// TIA Portal project "Oshop-Demo_v2" (V16)

(* hardware
DEVICE "ET 200SP-Station_1"  ET 200SP-Station
   slot 0: "Baugruppenträger_0"  Rack  6ES5 710-8MAx1
   slot 1: "PLC_1"  CPU 1512SP-1 PN  6ES7 512-1DK01-0AB0  V2.1
      slot 32768: "PROFINET-Schnittstelle_1"  X1
   slot 2: "DI 8x24VDC HF_1"  DI 8x24VDC HF  6ES7 131-6BF00-0CA0  V2.0
      slot 1: "DI 8x24VDC HF_1"  DI 8x24VDC HF
   slot 3: "CM 4xIO-Link_1"  CM 4xIO-Link  6ES7 137-6BD00-0BA0  V2.2
      slot 1: "CM 4xIO-Link_1"  6ES7 137-6BD00-0BA0
   slot 4: "DQ 8x24VDC/0.5A HF_1"  DQ 8x24VDC/0.5A HF  6ES7 132-6BF00-0CA0  V2.0
      slot 1: "DQ 8x24VDC/0.5A HF_1"  DQ 8x24VDC/0.5A HF
   slot 5: "Servermodul_1"  Server module  6ES7 193-6PA00-0AA0  V1.1
      slot 1: "Servermodul_1"  Server module
   slot 127: "BA 2xRJ45"  BA 2xRJ45  6ES7 193-6AR00-0AA0  V0.0
      slot 32769: "Port_1"  X1 P1  6ES7 193-6AR00-0AA0
      slot 32770: "Port_2"  X1 P2  6ES7 193-6AR00-0AA0
*)

// ===== PLC "PLC_1"  CPU 1512SP-1 PN =====

VAR_GLOBAL   // PLC tag table "Standard-Variablentabelle"
   "Tag_1" AT %IW102 : Word;
END_VAR

VAR_GLOBAL   // PLC tag table "IO-Link"
   "IOL-Hub_IN" AT %I100.0 : "udtIOL-Hub";
   "IOL-Hub_OUT" AT %Q100.0 : "udtIOL-Hub";
END_VAR

VAR_GLOBAL   // PLC tag table "DI"
   "Taster_Grün" AT %I0.0 : Bool;
   "Taster_WH_1" AT %I0.1 : Bool;
   "Taster_WH_2" AT %I0.2 : Bool;
END_VAR

VAR_GLOBAL   // PLC tag table "DO"
   "Lampe_WH_1" AT %Q0.1 : Bool;
   "Lampe_WH_2" AT %Q0.2 : Bool;
END_VAR

TYPE "udtToolCha_Sig_IN"
   STRUCT
      Tool_is_loaded : Bool;
      ToolStation_is_Locked : Bool;
      ToolStation_is_Released : Bool;
      ToolStation_is_Pos1 : Bool;
      ToolStation_is_Pos2 : Bool;
      ToolChanger_is_Locked : Bool;
      ToolChanger_is_Released : Bool;
      Lift_is_down : Bool;
      Lift_is_up : Bool;
   END_STRUCT;
END_TYPE

TYPE "udtToolCha_Sig_OUT"
   STRUCT
      ToolChanger : Bool;
      ToolStation_Select : Bool;
      ToolStation_Lock : Bool;
      Toolstation_Releas : Bool;
      Lift_down : Bool;
      Lift_up : Bool;
   END_STRUCT;
END_TYPE

TYPE "udtIOL-Hub"
   STRUCT
      "Byte" : Array[0..1] of Byte;
   END_STRUCT;
END_TYPE

DATA_BLOCK "Oshop_ToolChanger_DB"   // DB1
{ S7_Optimized_Access := 'TRUE' }
VERSION : 0.1
// stored: InstanceOfName Oshop_ToolChanger
"Oshop_ToolChanger"
BEGIN
END_DATA_BLOCK

DATA_BLOCK "GDB_Var"   // DB2
{ S7_Optimized_Access := 'TRUE' }
VERSION : 0.1
   VAR
      Tool : UInt;
   END_VAR
BEGIN
END_DATA_BLOCK

DATA_BLOCK "Tool_Select_DB"   // DB3
{ S7_Optimized_Access := 'TRUE' }
VERSION : 0.1
// stored: InstanceOfName Tool_Select
"Tool_Select"
BEGIN
END_DATA_BLOCK

FUNCTION_BLOCK "Oshop_ToolChanger"   // FB1, SCL
{ S7_Optimized_Access := 'TRUE' }
VERSION : 0.1
   VAR_INPUT
      Start : Bool;
      UseTool : UInt;
      P_Signals_IN : "udtToolCha_Sig_IN";
   END_VAR
   VAR_OUTPUT
      P_Signals_OUT : "udtToolCha_Sig_OUT";
   END_VAR
   VAR
      "Step" : UInt := 0;
      StepMem : UInt;
      StepDelay : TON_TIME;
      MeasuringTime : TON_TIME;
      RT_Start : R_TRIG;
   END_VAR
   VAR_TEMP
      InitPos : Bool;
   END_VAR
BEGIN
   (****************************************************************************************
    * program name:    Oshop_ToolChager
    * author:          ToSchi
    * owner:           Hochschule für Technik und Wirtschaft Dresden
    * 
    * description:
    * 
    * 
    * 
    * 
    ****************************************************************************************
    *)

   //trigger   -----------------------------------------------------------------------------
   #RT_Start(CLK := #Start);


   //timer   -------------------------------------------------------------------------------
   #MeasuringTime(IN := (#Step = 60),
                  PT := t#2s);

   #StepDelay(IN := (#Step = #StepMem),
              PT := t#2s);


   //initialization   ----------------------------------------------------------------------
   #InitPos := #P_Signals_IN.Lift_is_up AND #P_Signals_IN.ToolStation_is_Locked AND #P_Signals_IN.ToolChanger_is_Released;

   #StepMem := #Step;

   CASE #Step OF
       0:
           #P_Signals_OUT.Lift_down := 0;
           #P_Signals_OUT.Lift_up := 0;
           #P_Signals_OUT.ToolChanger := 0;
           #P_Signals_OUT.ToolStation_Lock := 0;
           #P_Signals_OUT.Toolstation_Releas := 0;
           #P_Signals_OUT.ToolStation_Select := 0;
           #Step := 1;


       1:
           #P_Signals_OUT.ToolStation_Lock := 1;
           #P_Signals_OUT.Toolstation_Releas := 0;
           IF #P_Signals_IN.ToolStation_is_Locked AND NOT #P_Signals_IN.ToolStation_is_Released AND #StepDelay.Q THEN
               #Step := 2;
           END_IF;


       2:
           #P_Signals_OUT.ToolChanger := 1;
           IF #P_Signals_IN.ToolChanger_is_Locked AND NOT #P_Signals_IN.ToolChanger_is_Released AND #StepDelay.Q THEN
               #Step := 3;
           END_IF;


       3:
           #P_Signals_OUT.ToolStation_Select := 0;
           IF #P_Signals_IN.ToolStation_is_Pos1 AND NOT #P_Signals_IN.ToolStation_is_Pos2 AND #StepDelay.Q THEN
               #Step := 4;
           END_IF;


       4:
           IF NOT #P_Signals_IN.Tool_is_loaded THEN
               #Step := 7;
           ELSE
               #Step := 5;
           END_IF;


       5:
           #P_Signals_OUT.ToolStation_Select := 1;
           IF NOT #P_Signals_IN.ToolStation_is_Pos1 AND #P_Signals_IN.ToolStation_is_Pos2 AND #StepDelay.Q THEN
               #Step := 6;
           END_IF;


       6:
           IF NOT #P_Signals_IN.Tool_is_loaded THEN
               #Step := 7;
           ELSE
               #Step := 9;
           END_IF;


       7:
           #P_Signals_OUT.ToolStation_Lock := 0;
           #P_Signals_OUT.Toolstation_Releas := 1;
           IF NOT #P_Signals_IN.ToolStation_is_Locked AND #P_Signals_IN.ToolStation_is_Released AND #StepDelay.Q THEN
               #Step := 9;
           END_IF;


       9:
           #P_Signals_OUT.Lift_up := 1;
           #P_Signals_OUT.Lift_down := 0;
           IF #P_Signals_IN.Lift_is_up AND NOT #P_Signals_IN.Lift_is_down AND #StepDelay.Q THEN
               #Step := 10;
           END_IF;


       10:
           #P_Signals_OUT.ToolStation_Lock := 1;
           #P_Signals_OUT.Toolstation_Releas := 0;
           IF #P_Signals_IN.ToolStation_is_Locked AND NOT #P_Signals_IN.ToolStation_is_Released AND #StepDelay.Q THEN
               #P_Signals_OUT.ToolChanger := 0;
               IF NOT #P_Signals_IN.ToolChanger_is_Locked AND #P_Signals_IN.ToolChanger_is_Released AND #StepDelay.Q THEN
                   #Step := 15;
               END_IF;
           END_IF;


       15:
           #P_Signals_OUT.Lift_up := TRUE;
           IF #InitPos AND #UseTool <> 0 AND #RT_Start.Q THEN
               #Step := #UseTool + 20;
           END_IF;


       21: 
           IF NOT #P_Signals_IN.ToolStation_is_Pos1 THEN
               #P_Signals_OUT.ToolStation_Select := 0;
           ELSE
               #Step := 25;
           END_IF;


       22: 
           IF NOT #P_Signals_IN.ToolStation_is_Pos2 THEN
               #P_Signals_OUT.ToolStation_Select := 1;
           ELSE
               #Step := 25;
           END_IF;


       25: 
           IF #P_Signals_IN.Tool_is_loaded THEN
               #Step := 30;
           ELSE
               //go to error step
               ;
           END_IF;


       30: 
           #P_Signals_OUT.ToolChanger := TRUE;

           IF #P_Signals_IN.ToolChanger_is_Locked THEN
               #Step := 40;
           END_IF;


       40:
           #P_Signals_OUT.ToolStation_Lock := FALSE;
           #P_Signals_OUT.Toolstation_Releas := TRUE;

           IF #P_Signals_IN.ToolStation_is_Released THEN
               #Step := 50;
           END_IF;


       50: 
           #P_Signals_OUT.Lift_up := FALSE;
           #P_Signals_OUT.Lift_down := TRUE;

           IF #P_Signals_IN.Lift_is_down THEN
               #Step := 60;
           END_IF;


       60:
           IF #MeasuringTime.Q THEN
               #Step := 70;
           END_IF;


       70:
           IF NOT #P_Signals_IN.Tool_is_loaded AND #P_Signals_IN.ToolStation_is_Released THEN
               #Step := 80;
           ELSE
               //go to error step
               ;
           END_IF;


       80: 
           #P_Signals_OUT.Lift_up := TRUE;
           #P_Signals_OUT.Lift_down := FALSE;

           IF #P_Signals_IN.Lift_is_up THEN
               #Step := 90;
           END_IF;


       90:
           #P_Signals_OUT.ToolStation_Lock := TRUE;
           #P_Signals_OUT.Toolstation_Releas := FALSE;

           IF #P_Signals_IN.ToolStation_is_Locked THEN
               #Step := 100;
           END_IF;


       100:
           #P_Signals_OUT.ToolChanger := FALSE;

           IF #P_Signals_IN.ToolChanger_is_Released THEN
               #Step := 15;
           END_IF;

   END_CASE;

   //---------------------------------------------------------------------------------------
   //End   ---------------------------------------------------------------------------------
END_FUNCTION_BLOCK

FUNCTION_BLOCK "Tool_Select"   // FB2, SCL
{ S7_Optimized_Access := 'TRUE' }
VERSION : 0.1
   VAR_INPUT
      Button_1 : Bool;
      Button_2 : Bool;
   END_VAR
   VAR_OUTPUT
      Lamp_1 : Bool;
      Lamp_2 : Bool;
      ToolNumber : UInt := 0;
   END_VAR
   VAR
      RT_Button_1 : R_TRIG;
      RT_Button_2 : R_TRIG;
   END_VAR
BEGIN
   (****************************************************************************************
    * program name:    ToolSelect
    * author:          ToSchi
    * owner:           Hochschule für Technik und Wirtschaft Dresden
    * 
    * description:
    * 
    * 
    * 
    * 
    ****************************************************************************************
    *)

   //trigger   -----------------------------------------------------------------------------
   #RT_Button_1(CLK := #Button_1);
   #RT_Button_2(CLK := #Button_2);


   //program   -----------------------------------------------------------------------------
   IF #RT_Button_1.Q THEN
       #ToolNumber := 1;
   ELSIF #RT_Button_2.Q THEN
       #ToolNumber := 2;
   ELSIF #RT_Button_1.Q AND #RT_Button_2.Q THEN
       #ToolNumber := 0;
   END_IF;

   #Lamp_1 := (#ToolNumber = 1);
   #Lamp_2 := (#ToolNumber = 2);

   //---------------------------------------------------------------------------------------
   //End   ---------------------------------------------------------------------------------
END_FUNCTION_BLOCK

ORGANIZATION_BLOCK "Main"   // OB1, LAD, ProgramCycle
TITLE = "Main Program Sweep (Cycle)"
{ S7_Optimized_Access := 'TRUE' }
VERSION : 0.1
   VAR_INPUT
      Initial_Call : Bool;   // Initial call of this OB
      Remanence : Bool;   // =True, if remanent data are available
   END_VAR
   VAR_TEMP
      Pos : DInt;
      RetVal : DInt;
      tmpByte : Byte;
   END_VAR
BEGIN

REGION Network 1
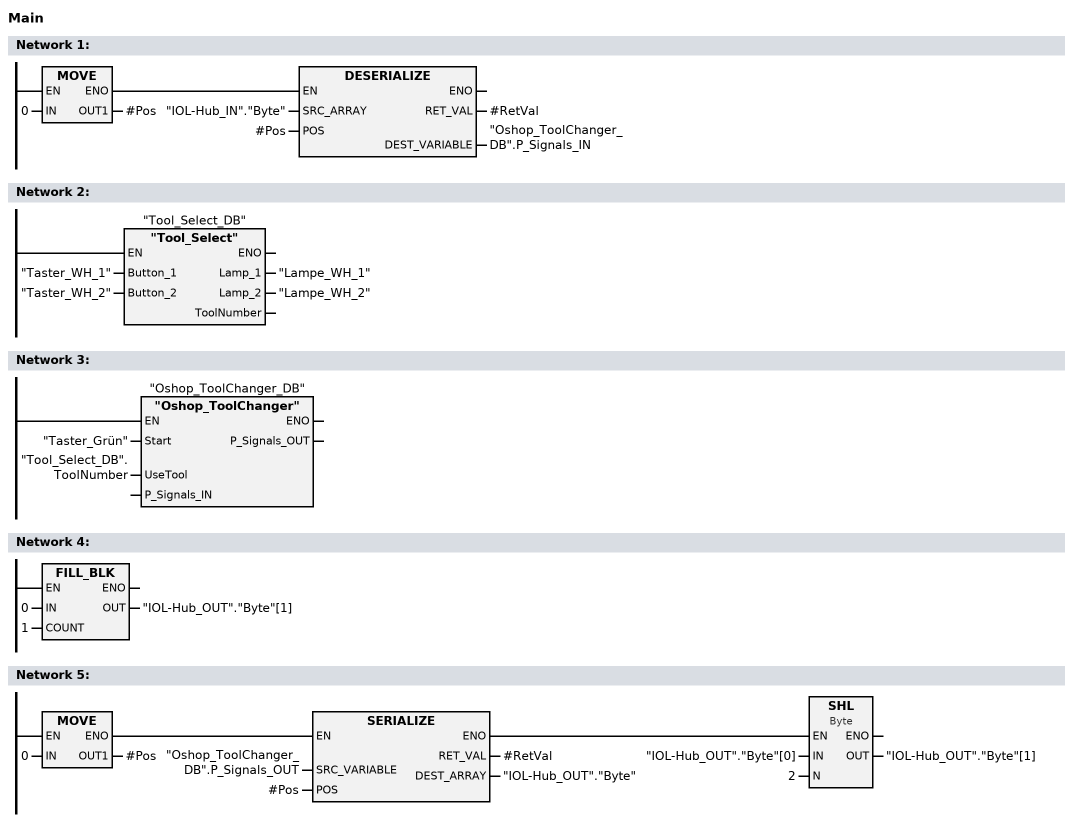
   // no SCL statement known for Deserialize: written as a call
   #Pos := 0;
   #RetVal := Deserialize(SRC_ARRAY := "IOL-Hub_IN"."Byte",
                          POS := #Pos,
                          DEST_VARIABLE => "Oshop_ToolChanger_DB".P_Signals_IN);
END_REGION

REGION Network 2
   RUNG wire#powerrail
      "Tool_Select_DB"(Button_1 := "Taster_WH_1", Button_2 := "Taster_WH_2", Lamp_1 => "Lampe_WH_1", Lamp_2 => "Lampe_WH_2", ToolNumber =>)
   END_RUNG
   // the same network as SCL:
   "Tool_Select_DB"(Button_1 := "Taster_WH_1",   // "Tool_Select"
                    Button_2 := "Taster_WH_2",
                    Lamp_1 => "Lampe_WH_1",
                    Lamp_2 => "Lampe_WH_2");
END_REGION

REGION Network 3
   RUNG wire#powerrail
      "Oshop_ToolChanger_DB"(Start := "Taster_Grün", UseTool := "Tool_Select_DB".ToolNumber, P_Signals_IN :=, P_Signals_OUT =>)
   END_RUNG
   // the same network as SCL:
   "Oshop_ToolChanger_DB"(Start := "Taster_Grün", UseTool := "Tool_Select_DB".ToolNumber);   // "Oshop_ToolChanger"
END_REGION

REGION Network 4
   RUNG wire#powerrail
      FillBlockI(in := 0, count := 1, out => "IOL-Hub_OUT"."Byte"[1])
   END_RUNG
   // the same network as SCL:
   FILL_BLK(IN := 0, COUNT := 1, OUT => "IOL-Hub_OUT"."Byte"[1]);
END_REGION

REGION Network 5
   // no SCL statement known for Serialize: written as a call
   // ENO of a box is taken as its EN; it also drops when the box reports an error
   #Pos := 0;
   #RetVal := Serialize(SRC_VARIABLE := "Oshop_ToolChanger_DB".P_Signals_OUT,
                        POS := #Pos,
                        DEST_ARRAY => "IOL-Hub_OUT"."Byte");
   "IOL-Hub_OUT"."Byte"[1] := SHL(IN := "IOL-Hub_OUT"."Byte"[0], N := 2);
END_REGION
END_ORGANIZATION_BLOCK

// ===== library: MasterCopy "ArrayOfByte_To_Word" =====

FUNCTION "ArrayOfByte_To_Word" : Void   // FC2, SCL
{ S7_Optimized_Access := 'TRUE' }
VERSION : 0.1
   VAR_INPUT
      Array_IN : Array[0..1] of Byte;
      StartPos : UInt;
   END_VAR
   VAR_OUTPUT
      Word_OUT : Word;
   END_VAR
BEGIN
   #Word_OUT := SHL_WORD(IN := #Word_OUT, N := #StartPos) OR #Array_IN[0];
END_FUNCTION

// ===== library: MasterCopy "Word_To_ArrayOfByte" =====

FUNCTION "Word_To_ArrayOfByte" : Void   // FC1, SCL
{ S7_Optimized_Access := 'TRUE' }
VERSION : 0.1
   VAR_INPUT
      Word_IN : Word;
   END_VAR
   VAR_OUTPUT
      Array_OUT : Array[0..1] of Byte;
   END_VAR
BEGIN
   #Array_OUT[1] := WORD_TO_BYTE(IN := #Word_IN);
   #Array_OUT[0] := WORD_TO_BYTE(IN := SHR_WORD(IN := #Word_IN, N := 8));
END_FUNCTION